                                   // Arc
                                   IF ((#statParameterValid.cmdParameters.circleParameters.arc AND #tempParseCounter = 1)
                                     OR (NOT #statParameterValid.cmdParameters.circleParameters.arc AND #tempParseCounter = 2))
                                     AND #statParameterDefinition.priorities.cmdParameters.circleParameters.arc > "LKINLANG_PRIO_UNRELEVANT"
                                   THEN
                                     // Get parameter value
                                     #tempParameterValue := #tempParsedValues.cmdParameters.circleParameters.arc;

                                     // Set Arc
                                     #statPathDataValue.valueLReal := #statActualCommand.pathDataElement.cmdParameters.circleParameters.arc;
                                     #statModalCmdValue.valueLReal := #statModalCommand.pathDataElement.cmdParameters.circleParameters.arc;
                                     #statModalPrgValue.valueLReal := #statModalProgram.pathDataElement.cmdParameters.circleParameters.arc;

                                     // Set value with follow val from above 
                                     #tempReturnVal := "LKinLang_SetValue"(parameterValue := #tempParameterValue,
                                                                           parameterPriority := #statParameterDefinition.priorities.cmdParameters.circleParameters.arc,
                                                                           validCountOfParameter := #statValidCounts.cmdParameters.circleParameters.arc,
                                                                           parameterValueMin := #MINVAL_LREAL,
                                                                           parameterValueMax := #MAXVAL_LREAL,
                                                                           properties := #statParameterDefinition.properties,
                                                                           errorString => #statErrorString,
                                                                           parameterCounter := #statElementCounter.cmdParameters.circleParameters.arc,
                                                                           priorityCounter := #statActualCommand.priority.cmdParameters.circleParameters.arc,
                                                                           modalCMDPrio := #statModalCommand.priority.cmdParameters.circleParameters.arc,
                                                                           modalPRGPrio := #statModalProgram.priority.cmdParameters.circleParameters.arc,
                                                                           parameterCounterInLine := #statElementCounterInLine.cmdParameters.circleParameters.arc,
                                                                           pathDataValue := #statPathDataValue,
                                                                           modalCMDPathDataValue := #statModalCmdValue,
                                                                           modalPRGPathDataValue := #statModalPrgValue);

                                     IF #tempReturnVal = 0 THEN
                                       #statActualCommand.pathDataElement.cmdParameters.circleParameters.arc := #statPathDataValue.valueLReal;
                                       #statModalCommand.pathDataElement.cmdParameters.circleParameters.arc := #statModalCmdValue.valueLReal;
                                       #statModalProgram.pathDataElement.cmdParameters.circleParameters.arc := #statModalPrgValue.valueLReal;
                                     ELSE
                                       // Error
                                       #statStatus := #ERR_PARSING;
                                       #statErrorString := CONCAT(IN1 := #statErrorString, IN2 := '; Line: ');
                                       #statErrorString := CONCAT(IN1 := #statErrorString, IN2 := UDINT_TO_STRING(#statTokenizedLine.lineNo));
                                       EXIT;
                                     END_IF;
                                   END_IF;


                                   // Radius
                                   IF (#statParameterValid.cmdParameters.circleParameters.radius AND #tempParseCounter = 1)
                                     OR (NOT #statParameterValid.cmdParameters.circleParameters.radius AND #tempParseCounter = 2)
                                     AND #statParameterDefinition.priorities.cmdParameters.circleParameters.radius > "LKINLANG_PRIO_UNRELEVANT"
                                   THEN
                                     // Get parameter value
                                     #tempParameterValue := #tempParsedValues.cmdParameters.circleParameters.radius;

                                     // Set Radius
                                     #statPathDataValue.valueLReal := #statActualCommand.pathDataElement.cmdParameters.circleParameters.radius;
                                     #statModalCmdValue.valueLReal := #statModalCommand.pathDataElement.cmdParameters.circleParameters.radius;
                                     #statModalPrgValue.valueLReal := #statModalProgram.pathDataElement.cmdParameters.circleParameters.radius;

                                     // Set value with follow val from above 
                                     #tempReturnVal := "LKinLang_SetValue"(parameterValue := #tempParameterValue,
                                                                           parameterPriority := #statParameterDefinition.priorities.cmdParameters.circleParameters.radius,
                                                                           validCountOfParameter := #statValidCounts.cmdParameters.circleParameters.radius,
                                                                           parameterValueMin := #MINVAL_LREAL,
                                                                           parameterValueMax := #MAXVAL_LREAL,
                                                                           properties := #statParameterDefinition.properties,
                                                                           errorString => #statErrorString,
                                                                           parameterCounter := #statElementCounter.cmdParameters.circleParameters.radius,
                                                                           priorityCounter := #statActualCommand.priority.cmdParameters.circleParameters.radius,
                                                                           modalCMDPrio := #statModalCommand.priority.cmdParameters.circleParameters.radius,
                                                                           modalPRGPrio := #statModalProgram.priority.cmdParameters.circleParameters.radius,
                                                                           parameterCounterInLine := #statElementCounterInLine.cmdParameters.circleParameters.radius,
                                                                           pathDataValue := #statPathDataValue,
                                                                           modalCMDPathDataValue := #statModalCmdValue,
                                                                           modalPRGPathDataValue := #statModalPrgValue);

                                     IF #tempReturnVal = 0 THEN
                                       #statActualCommand.pathDataElement.cmdParameters.circleParameters.radius := #statPathDataValue.valueLReal;
                                       #statModalCommand.pathDataElement.cmdParameters.circleParameters.radius := #statModalCmdValue.valueLReal;
                                       #statModalProgram.pathDataElement.cmdParameters.circleParameters.radius := #statModalPrgValue.valueLReal;
                                     ELSE
                                       // Error
                                       #statStatus := #ERR_PARSING;
                                       #statErrorString := CONCAT(IN1 := #statErrorString, IN2 := '; Line: ');
                                       #statErrorString := CONCAT(IN1 := #statErrorString, IN2 := UDINT_TO_STRING(#statTokenizedLine.lineNo));
                                       EXIT;
                                     END_IF;
                                   END_IF;

                                 END_IF;
                               END_REGION CIRCLE_PARAMETERS


                             END_IF;
                           END_REGION CMD_PARAMETERS

                           REGION BOOL_FLAGS
                             // In the first run the follow values are parsed
                             // If a flag was set in "GET_FOLLOW_VALUES" it is always written in the first index of "tempParsedValues"
                             // Direct values can be set in the complete array
                             // --> For each Flag which is set from follow values, increase the flag counter
                             // --> For each Flag which is set from direct values, increase the same flag counter
                             // Flag counter is only increased if flag is set but not for flagMode and remaining distance

                             // ----------------------------------------------------------------------------
                             // Set Flags
                             // ----------------------------------------------------------------------------
                             FOR #tempCounter := 1 TO "LKINCTRL_NO_OF_CMD_SETFLAGS" DO
                               IF (#statParameterValid.setFlags[#tempCounter].flag AND #tempParseCounter = 1)
                                 OR (#statParameterDefinition.directValues.setFlags[#tempCounter].flag <> #statParameterDefinitionEmpty.directValues.setFlags[#tempCounter].flag
                                 AND #tempParseCounter = 2)
                                 AND #statParameterDefinition.priorities.setFlags.flag > "LKINLANG_PRIO_UNRELEVANT"
                               THEN
                                 // Set actual flag number depending on counter
                                 #statActualFlagNumber := #statElementCounterInLine.setFlags.flag + #statElementCounter.setFlags.flag + 1;

                                 // Check flag index
                                 IF #statActualFlagNumber > "LKINCTRL_NO_OF_CMD_SETFLAGS" THEN
                                   // Error invalid flag index
                                   #statStatus := #ERR_PARSING;
                                   #statErrorString := CONCAT(IN1 := #statErrorString, IN2 := 'Only ');
                                   #statErrorString := CONCAT(IN1 := #statErrorString, IN2 := INT_TO_STRING("LKINCTRL_NO_OF_CMD_SETFLAGS"));
                                   #statErrorString := CONCAT(IN1 := #statErrorString, IN2 := ' Flags allowed per command');
                                   #statErrorString := CONCAT(IN1 := #statErrorString, IN2 := '; Line: ');
                                   #statErrorString := CONCAT(IN1 := #statErrorString, IN2 := UDINT_TO_STRING(#statTokenizedLine.lineNo));
                                   EXIT;
                                 ELSIF #statActualFlagNumber < 1 THEN
                                   // Error invalid flag index
                                   #statStatus := #ERR_PARSING;
                                   #statErrorString := CONCAT(IN1 := #statErrorString, IN2 := 'Invalid setflag index (<1) in line ');
                                   #statErrorString := CONCAT(IN1 := #statErrorString, IN2 := UDINT_TO_STRING(#statTokenizedLine.lineNo));
                                   EXIT;
                                 END_IF;

                                 // Get parameter value
                                 #tempParameterValue := #tempParsedValues.setFlags[#tempCounter].flag;

                                 #statPathDataValue.valueInt := #statActualCommand.pathDataElement.setFlags[#statActualFlagNumber].flag;
                                 #statModalCmdValue.valueInt := #statModalCommand.pathDataElement.setFlags[#statActualFlagNumber].flag;
                                 #statModalPrgValue.valueInt := #statModalProgram.pathDataElement.setFlags[#statActualFlagNumber].flag;

                                 // Set value with follow val from above 
                                 #tempReturnVal := "LKinLang_SetValue"(parameterValue := #tempParameterValue,
                                                                       parameterPriority := #statParameterDefinition.priorities.setFlags.flag,
                                                                       validCountOfParameter := #statValidCounts.setFlags.flag,
                                                                       parameterValueMin := -1,
                                                                       parameterValueMax := "LKINCTRL_NO_OF_LAST_SETFLAG",
                                                                       properties := #statParameterDefinition.properties,
                                                                       errorString => #statErrorString,
                                                                       parameterCounter := #statElementCounter.setFlags.flag,
                                                                       priorityCounter := #statActualCommand.priority.setFlags[#statActualFlagNumber].flag,
                                                                       modalCMDPrio := #statModalCommand.priority.setFlags[#statActualFlagNumber].flag,
                                                                       modalPRGPrio := #statModalProgram.priority.setFlags[#statActualFlagNumber].flag,
                                                                       parameterCounterInLine := #statElementCounterInLine.setFlags.flag,
                                                                       pathDataValue := #statPathDataValue,
                                                                       modalCMDPathDataValue := #statModalCmdValue,
                                                                       modalPRGPathDataValue := #statModalPrgValue);

                                 IF #tempReturnVal = 0 THEN // Parameter is ok
                                   #statActualCommand.pathDataElement.setFlags[#statActualFlagNumber].flag := #statPathDataValue.valueInt;
                                   #statModalCommand.pathDataElement.setFlags[#statActualFlagNumber].flag := #statModalCmdValue.valueInt;
                                   #statModalProgram.pathDataElement.setFlags[#statActualFlagNumber].flag := #statModalPrgValue.valueInt;
                                 ELSE
                                   // Error
                                   #statStatus := #ERR_PARSING;
                                   #statErrorString := CONCAT(IN1 := #statErrorString, IN2 := '; Line: ');
                                   #statErrorString := CONCAT(IN1 := #statErrorString, IN2 := UDINT_TO_STRING(#statTokenizedLine.lineNo));
                                   EXIT;
                                 END_IF;
                               END_IF;

                               // ----------------------------------------------------------------------------
                               // Flag Mode
                               // ----------------------------------------------------------------------------
                               IF (#statParameterValid.setFlags[#tempCounter].flagMode AND #tempParseCounter = 1)
                                 OR (#statParameterDefinition.directValues.setFlags[#tempCounter].flagMode <> #statParameterDefinitionEmpty.directValues.setFlags[#tempCounter].flagMode
                                 AND #tempParseCounter = 2)
                                 AND #statParameterDefinition.priorities.setFlags.flagMode > "LKINLANG_PRIO_UNRELEVANT"
                               THEN
                                 // Set actual flag number depending on counter
                                 #statActualFlagNumber := #statElementCounterInLine.setFlags.flagMode + #statElementCounter.setFlags.flagMode + 1;

                                 // Check flag index
                                 IF #statActualFlagNumber > "LKINCTRL_NO_OF_CMD_SETFLAGS" THEN
                                   // Error invalid flag index
                                   #statStatus := #ERR_PARSING;
                                   #statErrorString := CONCAT(IN1 := #statErrorString, IN2 := 'Only ');
                                   #statErrorString := CONCAT(IN1 := #statErrorString, IN2 := INT_TO_STRING("LKINCTRL_NO_OF_CMD_SETFLAGS"));
                                   #statErrorString := CONCAT(IN1 := #statErrorString, IN2 := ' Flags allowed per command');
                                   #statErrorString := CONCAT(IN1 := #statErrorString, IN2 := '; Line: ');
                                   #statErrorString := CONCAT(IN1 := #statErrorString, IN2 := UDINT_TO_STRING(#statTokenizedLine.lineNo));
                                   EXIT;
                                 ELSIF #statActualFlagNumber < 1 THEN
                                   // Error invalid flag index
                                   #statStatus := #ERR_PARSING;
                                   #statErrorString := CONCAT(IN1 := #statErrorString, IN2 := 'Invalid setflag index (<1) in line ');
                                   #statErrorString := CONCAT(IN1 := #statErrorString, IN2 := UDINT_TO_STRING(#statTokenizedLine.lineNo));
                                   EXIT;
                                 END_IF;

                                 // Get parameter value
                                 #tempParameterValue := #tempParsedValues.setFlags[#tempCounter].flagMode;

                                 #statPathDataValue.valueInt := #statActualCommand.pathDataElement.setFlags[#statActualFlagNumber].flagMode;
                                 #statModalCmdValue.valueInt := #statModalCommand.pathDataElement.setFlags[#statActualFlagNumber].flagMode;
                                 #statModalPrgValue.valueInt := #statModalProgram.pathDataElement.setFlags[#statActualFlagNumber].flagMode;

                                 // Set value with follow val from above 
                                 #tempReturnVal := "LKinLang_SetValue"(parameterValue := #tempParameterValue,
                                                                       parameterPriority := #statParameterDefinition.priorities.setFlags.flagMode,
                                                                       validCountOfParameter := #statValidCounts.setFlags.flagMode,
                                                                       parameterValueMin := 0,
                                                                       parameterValueMax := 15,
                                                                       properties := #statParameterDefinition.properties,
                                                                       errorString => #statErrorString,
                                                                       parameterCounter := #statElementCounter.setFlags.flagMode,
                                                                       priorityCounter := #statActualCommand.priority.setFlags[#statActualFlagNumber].flagMode,
                                                                       modalCMDPrio := #statModalCommand.priority.setFlags[#statActualFlagNumber].flagMode,
                                                                       modalPRGPrio := #statModalProgram.priority.setFlags[#statActualFlagNumber].flagMode,
                                                                       parameterCounterInLine := #statElementCounterInLine.setFlags.flagMode,
                                                                       pathDataValue := #statPathDataValue,
                                                                       modalCMDPathDataValue := #statModalCmdValue,
                                                                       modalPRGPathDataValue := #statModalPrgValue);

                                 IF #tempReturnVal = 0 THEN // Parameter is ok
                                   #statActualCommand.pathDataElement.setFlags[#statActualFlagNumber].flagMode := INT_TO_USINT(#statPathDataValue.valueInt);
                                   #statModalCommand.pathDataElement.setFlags[#statActualFlagNumber].flagMode := INT_TO_USINT(#statModalCmdValue.valueInt);
                                   #statModalProgram.pathDataElement.setFlags[#statActualFlagNumber].flagMode := INT_TO_USINT(#statModalPrgValue.valueInt);
                                 ELSE
                                   // Error
                                   #statStatus := #ERR_PARSING;
                                   #statErrorString := CONCAT(IN1 := #statErrorString, IN2 := '; Line: ');
                                   #statErrorString := CONCAT(IN1 := #statErrorString, IN2 := UDINT_TO_STRING(#statTokenizedLine.lineNo));
                                   EXIT;
                                 END_IF;
                               END_IF;


                               // ----------------------------------------------------------------------------
                               // Remaining Distance
                               // ----------------------------------------------------------------------------
                               IF (#statParameterValid.setFlags[#tempCounter].remainingDistance AND #tempParseCounter = 1)
                                 OR (#statParameterDefinition.directValues.setFlags[#tempCounter].remainingDistance <> #statParameterDefinitionEmpty.directValues.setFlags[#tempCounter].remainingDistance
                                 AND #tempParseCounter = 2)
                                 AND #statParameterDefinition.priorities.setFlags.remainingDistance > "LKINLANG_PRIO_UNRELEVANT"
                               THEN
                                 // Set actual flag number depending on counter
                                 #statActualFlagNumber := #statElementCounterInLine.setFlags.remainingDistance + #statElementCounter.setFlags.remainingDistance + 1;

                                 // Check flag index
                                 IF #statActualFlagNumber > "LKINCTRL_NO_OF_CMD_SETFLAGS" THEN
                                   // Error invalid flag index
                                   #statStatus := #ERR_PARSING;
                                   #statErrorString := CONCAT(IN1 := #statErrorString, IN2 := 'Only ');
                                   #statErrorString := CONCAT(IN1 := #statErrorString, IN2 := INT_TO_STRING("LKINCTRL_NO_OF_CMD_SETFLAGS"));
                                   #statErrorString := CONCAT(IN1 := #statErrorString, IN2 := ' Flags allowed per command');
                                   #statErrorString := CONCAT(IN1 := #statErrorString, IN2 := '; Line: ');
                                   #statErrorString := CONCAT(IN1 := #statErrorString, IN2 := UDINT_TO_STRING(#statTokenizedLine.lineNo));
                                   EXIT;
                                 ELSIF #statActualFlagNumber < 1 THEN
                                   // Error invalid flag index
                                   #statStatus := #ERR_PARSING;
                                   #statErrorString := CONCAT(IN1 := #statErrorString, IN2 := 'Invalid setflag index (<1) in line ');
                                   #statErrorString := CONCAT(IN1 := #statErrorString, IN2 := UDINT_TO_STRING(#statTokenizedLine.lineNo));
                                   EXIT;
                                 END_IF;

                                 // Get parameter value
                                 #tempParameterValue := #tempParsedValues.setFlags[#tempCounter].remainingDistance;

                                 #statPathDataValue.valueLReal := #statActualCommand.pathDataElement.setFlags[#statActualFlagNumber].remainingDistance;
                                 #statModalCmdValue.valueLReal := #statModalCommand.pathDataElement.setFlags[#statActualFlagNumber].remainingDistance;
                                 #statModalPrgValue.valueLReal := #statModalProgram.pathDataElement.setFlags[#statActualFlagNumber].remainingDistance;

                                 // Set value with follow val from above 
                                 #tempReturnVal := "LKinLang_SetValue"(parameterValue := #tempParameterValue,
                                                                       parameterPriority := #statParameterDefinition.priorities.setFlags.remainingDistance,
                                                                       validCountOfParameter := #statValidCounts.setFlags.remainingDistance,
                                                                       parameterValueMin := #MINVAL_LREAL,
                                                                       parameterValueMax := #MAXVAL_LREAL,
                                                                       properties := #statParameterDefinition.properties,
                                                                       errorString => #statErrorString,
                                                                       parameterCounter := #statElementCounter.setFlags.remainingDistance,
                                                                       priorityCounter := #statActualCommand.priority.setFlags[#statActualFlagNumber].remainingDistance,
                                                                       modalCMDPrio := #statModalCommand.priority.setFlags[#statActualFlagNumber].remainingDistance,
                                                                       modalPRGPrio := #statModalProgram.priority.setFlags[#statActualFlagNumber].remainingDistance,
                                                                       parameterCounterInLine := #statElementCounterInLine.setFlags.remainingDistance,
                                                                       pathDataValue := #statPathDataValue,
                                                                       modalCMDPathDataValue := #statModalCmdValue,
                                                                       modalPRGPathDataValue := #statModalPrgValue);

                                 IF #tempReturnVal = 0 THEN // Parameter is ok
                                   #statActualCommand.pathDataElement.setFlags[#statActualFlagNumber].remainingDistance := #statPathDataValue.valueLReal;
                                   #statModalCommand.pathDataElement.setFlags[#statActualFlagNumber].remainingDistance := #statModalCmdValue.valueLReal;
                                   #statModalProgram.pathDataElement.setFlags[#statActualFlagNumber].remainingDistance := #statModalPrgValue.valueLReal;
                                 ELSE
                                   // Error
                                   #statStatus := #ERR_PARSING;
                                   #statErrorString := CONCAT(IN1 := #statErrorString, IN2 := '; Line: ');
                                   #statErrorString := CONCAT(IN1 := #statErrorString, IN2 := UDINT_TO_STRING(#statTokenizedLine.lineNo));
                                   EXIT;
                                 END_IF;
                               END_IF;

                             END_FOR;
                           END_REGION BOOL_FLAGS

                           REGION LREAL_FLAGS
                             // ----------------------------------------------------------------------------
                             // Set LREAL Flags
                             // ----------------------------------------------------------------------------
                             FOR #tempCounter := 1 TO "LKINCTRL_NO_OF_CMD_VALUEFLAGS" DO
                               IF (#statParameterValid.valueFlags[#tempCounter].flag AND #tempParseCounter = 1)
                                 OR (#statParameterDefinition.directValues.valueFlags[#tempCounter].flag <> #statParameterDefinitionEmpty.directValues.valueFlags[#tempCounter].flag
                                 AND #tempParseCounter = 2)
                                 AND #statParameterDefinition.priorities.valueFlags.flag > "LKINLANG_PRIO_UNRELEVANT"
                               THEN
                                 // Set actual flag number depending on counter
                                 #statActualValueFlagNumber := #statElementCounterInLine.valueFlags.flag + #statElementCounter.valueFlags.flag + 1;

                                 // Check flag index
                                 IF #statActualValueFlagNumber > "LKINCTRL_NO_OF_CMD_VALUEFLAGS" THEN
                                   // Error
                                   #statStatus := #ERR_PARSING;
                                   #statErrorString := CONCAT(IN1 := #statErrorString, IN2 := 'Only ');
                                   #statErrorString := CONCAT(IN1 := #statErrorString, IN2 := INT_TO_STRING("LKINCTRL_NO_OF_CMD_VALUEFLAGS"));
                                   #statErrorString := CONCAT(IN1 := #statErrorString, IN2 := ' Flags allowed per command');
                                   #statErrorString := CONCAT(IN1 := #statErrorString, IN2 := '; Line: ');
                                   #statErrorString := CONCAT(IN1 := #statErrorString, IN2 := UDINT_TO_STRING(#statTokenizedLine.lineNo));
                                   EXIT;
                                 ELSIF #statActualValueFlagNumber < 1 THEN
                                   // Error invalid flag index
                                   #statStatus := #ERR_PARSING;
                                   #statErrorString := CONCAT(IN1 := #statErrorString, IN2 := 'Invalid valueflag index (<1) in line ');
                                   #statErrorString := CONCAT(IN1 := #statErrorString, IN2 := UDINT_TO_STRING(#statTokenizedLine.lineNo));
                                   EXIT;
                                 END_IF;

                                 // Get parameter value
                                 #tempParameterValue := #tempParsedValues.valueFlags[#tempCounter].flag;

                                 #statPathDataValue.valueInt := #statActualCommand.pathDataElement.valueFlags[#statActualValueFlagNumber].flag;
                                 #statModalCmdValue.valueInt := #statModalCommand.pathDataElement.valueFlags[#statActualValueFlagNumber].flag;
                                 #statModalPrgValue.valueInt := #statModalProgram.pathDataElement.valueFlags[#statActualValueFlagNumber].flag;

                                 // Set value with follow val from above 
                                 #tempReturnVal := "LKinLang_SetValue"(parameterValue := #tempParameterValue,
                                                                       parameterPriority := #statParameterDefinition.priorities.valueFlags.flag,
                                                                       validCountOfParameter := #statValidCounts.valueFlags.flag,
                                                                       parameterValueMin := -1,
                                                                       parameterValueMax := "LKINCTRL_NO_OF_LAST_VALUEFLAG",
                                                                       properties := #statParameterDefinition.properties,
                                                                       errorString => #statErrorString,
                                                                       parameterCounter := #statElementCounter.valueFlags.flag,
                                                                       priorityCounter := #statActualCommand.priority.valueFlags[#statActualValueFlagNumber].flag,
                                                                       modalCMDPrio := #statModalCommand.priority.valueFlags[#statActualValueFlagNumber].flag,
                                                                       modalPRGPrio := #statModalProgram.priority.valueFlags[#statActualValueFlagNumber].flag,
                                                                       parameterCounterInLine := #statElementCounterInLine.valueFlags.flag,
                                                                       pathDataValue := #statPathDataValue,
                                                                       modalCMDPathDataValue := #statModalCmdValue,
                                                                       modalPRGPathDataValue := #statModalPrgValue);

                                 IF #tempReturnVal = 0 THEN // Parameter is ok
                                   #statActualCommand.pathDataElement.valueFlags[#statActualValueFlagNumber].flag := #statPathDataValue.valueInt;
                                   #statModalCommand.pathDataElement.valueFlags[#statActualValueFlagNumber].flag := #statModalCmdValue.valueInt;
                                   #statModalProgram.pathDataElement.valueFlags[#statActualValueFlagNumber].flag := #statModalPrgValue.valueInt;
                                 ELSE
                                   // Error
                                   #statStatus := #ERR_PARSING;
                                   #statErrorString := CONCAT(IN1 := #statErrorString, IN2 := '; Line: ');
                                   #statErrorString := CONCAT(IN1 := #statErrorString, IN2 := UDINT_TO_STRING(#statTokenizedLine.lineNo));
                                   EXIT;
                                 END_IF;
                               END_IF;

                               // ----------------------------------------------------------------------------
                               // Flag Value
                               // ----------------------------------------------------------------------------
                               IF (#statParameterValid.valueFlags[#tempCounter].value AND #tempParseCounter = 1)
                                 OR (#statParameterDefinition.directValues.valueFlags[#tempCounter].value <> #statParameterDefinitionEmpty.directValues.valueFlags[#tempCounter].value
                                 AND #tempParseCounter = 2)
                                 AND #statParameterDefinition.priorities.valueFlags.value > "LKINLANG_PRIO_UNRELEVANT"
                               THEN
                                 // Set actual flag number depending on counter
                                 #statActualValueFlagNumber := #statElementCounterInLine.valueFlags.value + #statElementCounter.valueFlags.value + 1;

                                 // Check flag index
                                 IF #statActualValueFlagNumber > "LKINCTRL_NO_OF_CMD_VALUEFLAGS" THEN
                                   // Error
                                   #statStatus := #ERR_PARSING;
                                   #statErrorString := CONCAT(IN1 := #statErrorString, IN2 := 'Only ');
                                   #statErrorString := CONCAT(IN1 := #statErrorString, IN2 := INT_TO_STRING("LKINCTRL_NO_OF_CMD_VALUEFLAGS"));
                                   #statErrorString := CONCAT(IN1 := #statErrorString, IN2 := ' Flags allowed per command');
                                   #statErrorString := CONCAT(IN1 := #statErrorString, IN2 := '; Line: ');
                                   #statErrorString := CONCAT(IN1 := #statErrorString, IN2 := UDINT_TO_STRING(#statTokenizedLine.lineNo));
                                   EXIT;
                                 ELSIF #statActualValueFlagNumber < 1 THEN
                                   // Error invalid flag index
                                   #statStatus := #ERR_PARSING;
                                   #statErrorString := CONCAT(IN1 := #statErrorString, IN2 := 'Invalid valueflag index (<1) in line ');
                                   #statErrorString := CONCAT(IN1 := #statErrorString, IN2 := UDINT_TO_STRING(#statTokenizedLine.lineNo));
                                   EXIT;
                                 END_IF;

                                 // Get parameter value
                                 #tempParameterValue := #tempParsedValues.valueFlags[#tempCounter].value;

                                 #statPathDataValue.valueLReal := #statActualCommand.pathDataElement.valueFlags[#statActualValueFlagNumber].value;
                                 #statModalCmdValue.valueLReal := #statModalCommand.pathDataElement.valueFlags[#statActualValueFlagNumber].value;
                                 #statModalPrgValue.valueLReal := #statModalProgram.pathDataElement.valueFlags[#statActualValueFlagNumber].value;

                                 // Set value with follow val from above 
                                 #tempReturnVal := "LKinLang_SetValue"(parameterValue := #tempParameterValue,
                                                                       parameterPriority := #statParameterDefinition.priorities.valueFlags.value,
                                                                       validCountOfParameter := #statValidCounts.valueFlags.value,
                                                                       parameterValueMin := #MINVAL_LREAL,
                                                                       parameterValueMax := #MAXVAL_LREAL,
                                                                       properties := #statParameterDefinition.properties,
                                                                       errorString => #statErrorString,
                                                                       parameterCounter := #statElementCounter.valueFlags.value,
                                                                       priorityCounter := #statActualCommand.priority.valueFlags[#statActualValueFlagNumber].value,
                                                                       modalCMDPrio := #statModalCommand.priority.valueFlags[#statActualValueFlagNumber].value,
                                                                       modalPRGPrio := #statModalProgram.priority.valueFlags[#statActualValueFlagNumber].value,
                                                                       parameterCounterInLine := #statElementCounterInLine.valueFlags.value,
                                                                       pathDataValue := #statPathDataValue,
                                                                       modalCMDPathDataValue := #statModalCmdValue,
                                                                       modalPRGPathDataValue := #statModalPrgValue);

                                 IF #tempReturnVal = 0 THEN // Parameter is ok
                                   #statActualCommand.pathDataElement.valueFlags[#statActualValueFlagNumber].value := #statPathDataValue.valueLReal;
                                   #statModalCommand.pathDataElement.valueFlags[#statActualValueFlagNumber].value := #statModalCmdValue.valueLReal;
                                   #statModalProgram.pathDataElement.valueFlags[#statActualValueFlagNumber].value := #statModalPrgValue.valueLReal;
                                 ELSE
                                   // Error
                                   #statStatus := #ERR_PARSING;
                                   #statErrorString := CONCAT(IN1 := #statErrorString, IN2 := '; Line: ');
                                   #statErrorString := CONCAT(IN1 := #statErrorString, IN2 := UDINT_TO_STRING(#statTokenizedLine.lineNo));
                                   EXIT;
                                 END_IF;
                               END_IF;

                               // ----------------------------------------------------------------------------
                               // Flag Mode
                               // ----------------------------------------------------------------------------
                               IF (#statParameterValid.valueFlags[#tempCounter].flagMode AND #tempParseCounter = 1)
                                 OR (#statParameterDefinition.directValues.valueFlags[#tempCounter].flagMode <> #statParameterDefinitionEmpty.directValues.valueFlags[#tempCounter].flagMode
                                 AND #tempParseCounter = 2)
                                 AND #statParameterDefinition.priorities.valueFlags.flagMode > "LKINLANG_PRIO_UNRELEVANT"
                               THEN
                                 // Set actual flag number depending on counter
                                 #statActualValueFlagNumber := #statElementCounterInLine.valueFlags.flagMode + #statElementCounter.valueFlags.flagMode + 1;

                                 // Check flag index
                                 IF #statActualValueFlagNumber > "LKINCTRL_NO_OF_CMD_VALUEFLAGS" THEN
                                   // Error
                                   #statStatus := #ERR_PARSING;
                                   #statErrorString := CONCAT(IN1 := #statErrorString, IN2 := 'Only ');
                                   #statErrorString := CONCAT(IN1 := #statErrorString, IN2 := INT_TO_STRING("LKINCTRL_NO_OF_CMD_VALUEFLAGS"));
                                   #statErrorString := CONCAT(IN1 := #statErrorString, IN2 := ' Flags allowed per command');
                                   #statErrorString := CONCAT(IN1 := #statErrorString, IN2 := '; Line: ');
                                   #statErrorString := CONCAT(IN1 := #statErrorString, IN2 := UDINT_TO_STRING(#statTokenizedLine.lineNo));
                                   EXIT;
                                 ELSIF #statActualValueFlagNumber < 1 THEN
                                   // Error invalid flag index
                                   #statStatus := #ERR_PARSING;
                                   #statErrorString := CONCAT(IN1 := #statErrorString, IN2 := 'Invalid valueflag index (<1) in line ');
                                   #statErrorString := CONCAT(IN1 := #statErrorString, IN2 := UDINT_TO_STRING(#statTokenizedLine.lineNo));
                                   EXIT;
                                 END_IF;

                                 // Get parameter value
                                 #tempParameterValue := #tempParsedValues.valueFlags[#tempCounter].flagMode;

                                 #statPathDataValue.valueInt := #statActualCommand.pathDataElement.valueFlags[#statActualValueFlagNumber].flagMode;
                                 #statModalCmdValue.valueInt := #statModalCommand.pathDataElement.valueFlags[#statActualValueFlagNumber].flagMode;
                                 #statModalPrgValue.valueInt := #statModalProgram.pathDataElement.valueFlags[#statActualValueFlagNumber].flagMode;

                                 // Set value with follow val from above 
                                 #tempReturnVal := "LKinLang_SetValue"(parameterValue := #tempParameterValue,
                                                                       parameterPriority := #statParameterDefinition.priorities.valueFlags.flagMode,
                                                                       validCountOfParameter := #statValidCounts.valueFlags.flagMode,
                                                                       parameterValueMin := 0,
                                                                       parameterValueMax := 15,
                                                                       properties := #statParameterDefinition.properties,
                                                                       errorString => #statErrorString,
                                                                       parameterCounter := #statElementCounter.valueFlags.flagMode,
                                                                       priorityCounter := #statActualCommand.priority.valueFlags[#statActualValueFlagNumber].flagMode,
                                                                       modalCMDPrio := #statModalCommand.priority.valueFlags[#statActualValueFlagNumber].flagMode,
                                                                       modalPRGPrio := #statModalProgram.priority.valueFlags[#statActualValueFlagNumber].flagMode,
                                                                       parameterCounterInLine := #statElementCounterInLine.valueFlags.flagMode,
                                                                       pathDataValue := #statPathDataValue,
                                                                       modalCMDPathDataValue := #statModalCmdValue,
                                                                       modalPRGPathDataValue := #statModalPrgValue);

                                 IF #tempReturnVal = 0 THEN // Parameter is ok
                                   #statActualCommand.pathDataElement.valueFlags[#statActualValueFlagNumber].flagMode := INT_TO_USINT(#statPathDataValue.valueInt);
                                   #statModalCommand.pathDataElement.valueFlags[#statActualValueFlagNumber].flagMode := INT_TO_USINT(#statModalCmdValue.valueInt);
                                   #statModalProgram.pathDataElement.valueFlags[#statActualValueFlagNumber].flagMode := INT_TO_USINT(#statModalPrgValue.valueInt);
                                 ELSE
                                   // Error
                                   #statStatus := #ERR_PARSING;
                                   #statErrorString := CONCAT(IN1 := #statErrorString, IN2 := '; Line: ');
                                   #statErrorString := CONCAT(IN1 := #statErrorString, IN2 := UDINT_TO_STRING(#statTokenizedLine.lineNo));
                                   EXIT;
                                 END_IF;
                               END_IF;


                               // ----------------------------------------------------------------------------
                               // Remaining Distance
                               // ----------------------------------------------------------------------------
                               IF (#statParameterValid.valueFlags[#tempCounter].remainingDistance AND #tempParseCounter = 1)
                                 OR (#statParameterDefinition.directValues.valueFlags[#tempCounter].remainingDistance <> #statParameterDefinitionEmpty.directValues.valueFlags[#tempCounter].remainingDistance
                                 AND #tempParseCounter = 2)
                                 AND #statParameterDefinition.priorities.valueFlags.remainingDistance > "LKINLANG_PRIO_UNRELEVANT"
                               THEN
                                 // Set actual flag number depending on counter
                                 #statActualValueFlagNumber := #statElementCounterInLine.valueFlags.remainingDistance + #statElementCounter.valueFlags.remainingDistance + 1;

                                 // Check flag index
                                 IF #statActualValueFlagNumber > "LKINCTRL_NO_OF_CMD_VALUEFLAGS" THEN
                                   // Error
                                   #statStatus := #ERR_PARSING;
                                   #statErrorString := CONCAT(IN1 := #statErrorString, IN2 := 'Only ');
                                   #statErrorString := CONCAT(IN1 := #statErrorString, IN2 := INT_TO_STRING("LKINCTRL_NO_OF_CMD_VALUEFLAGS"));
                                   #statErrorString := CONCAT(IN1 := #statErrorString, IN2 := ' Flags allowed per command');
                                   #statErrorString := CONCAT(IN1 := #statErrorString, IN2 := '; Line: ');
                                   #statErrorString := CONCAT(IN1 := #statErrorString, IN2 := UDINT_TO_STRING(#statTokenizedLine.lineNo));
                                   EXIT;
                                 ELSIF #statActualValueFlagNumber < 1 THEN
                                   // Error invalid flag index
                                   #statStatus := #ERR_PARSING;
                                   #statErrorString := CONCAT(IN1 := #statErrorString, IN2 := 'Invalid valueflag index (<1) in line ');
                                   #statErrorString := CONCAT(IN1 := #statErrorString, IN2 := UDINT_TO_STRING(#statTokenizedLine.lineNo));
                                   EXIT;
                                 END_IF;

                                 // Get parameter value
                                 #tempParameterValue := #tempParsedValues.valueFlags[#tempCounter].remainingDistance;

                                 #statPathDataValue.valueLReal := #statActualCommand.pathDataElement.valueFlags[#statActualValueFlagNumber].remainingDistance;
                                 #statModalCmdValue.valueLReal := #statModalCommand.pathDataElement.valueFlags[#statActualValueFlagNumber].remainingDistance;
                                 #statModalPrgValue.valueLReal := #statModalProgram.pathDataElement.valueFlags[#statActualValueFlagNumber].remainingDistance;